   		OWF_Add_c.10:=OWF_Result[10].31;
   		OWF_Result[10].31:=0;
   		OWF_Result[11]:=OWF_Result[11] + 742245961+OWF_Add_c;
   		OWF_Add_c.11:=OWF_Result[11].31;
   		OWF_Result[11].31:=0;
   		OWF_Result[12]:=OWF_Result[12] + 1527470677+OWF_Add_c;
   		OWF_Add_c.12:=OWF_Result[12].31;
   		OWF_Result[12].31:=0;
   		OWF_Result[13]:=OWF_Result[13] + 104891933+OWF_Add_c;
   		OWF_Add_c.13:=OWF_Result[13].31;
   		OWF_Result[13].31:=0;
   		OWF_Result[14]:=OWF_Result[14] + 1414596320+OWF_Add_c;
   		OWF_Add_c.14:=OWF_Result[14].31;
   		OWF_Result[14].31:=0;
   		OWF_Result[15]:=OWF_Result[15] + 848151661+OWF_Add_c;
   		OWF_Add_c.15:=OWF_Result[15].31;
   		OWF_Result[15].31:=0;
   		OWF_Result[16]:=OWF_Result[16] + 1988122072+OWF_Add_c;
   		OWF_Add_c.16:=OWF_Result[16].31;
   		OWF_Result[16].31:=0;
   	End_If;
   	If OWF_Input[10].[29] Then
   		OWF_Result[0]:=OWF_Result[0] + 197995467+OWF_Add_c;
   		OWF_Add_c.0:=OWF_Result[0].31;
   		OWF_Result[0].31:=0;
   		OWF_Result[1]:=OWF_Result[1] + 1401962007+OWF_Add_c;
   		OWF_Add_c.1:=OWF_Result[1].31;
   		OWF_Result[1].31:=0;
   		OWF_Result[2]:=OWF_Result[2] + 1030218683+OWF_Add_c;
   		OWF_Add_c.2:=OWF_Result[2].31;
   		OWF_Result[2].31:=0;
   		OWF_Result[3]:=OWF_Result[3] + 1917186559+OWF_Add_c;
   		OWF_Add_c.3:=OWF_Result[3].31;
   		OWF_Result[3].31:=0;
   		OWF_Result[4]:=OWF_Result[4] + 1642815876+OWF_Add_c;
   		OWF_Add_c.4:=OWF_Result[4].31;
   		OWF_Result[4].31:=0;
   		OWF_Result[5]:=OWF_Result[5] + 126047613+OWF_Add_c;
   		OWF_Add_c.5:=OWF_Result[5].31;
   		OWF_Result[5].31:=0;
   		OWF_Result[6]:=OWF_Result[6] + 559790140+OWF_Add_c;
   		OWF_Add_c.6:=OWF_Result[6].31;
   		OWF_Result[6].31:=0;
   		OWF_Result[7]:=OWF_Result[7] + 2038093848+OWF_Add_c;
   		OWF_Add_c.7:=OWF_Result[7].31;
   		OWF_Result[7].31:=0;
   		OWF_Result[8]:=OWF_Result[8] + 221043685+OWF_Add_c;
   		OWF_Add_c.8:=OWF_Result[8].31;
   		OWF_Result[8].31:=0;
   		OWF_Result[9]:=OWF_Result[9] + 1671325631+OWF_Add_c;
   		OWF_Add_c.9:=OWF_Result[9].31;
   		OWF_Result[9].31:=0;
   		OWF_Result[10]:=OWF_Result[10] + 466139389+OWF_Add_c;
   		OWF_Add_c.10:=OWF_Result[10].31;
   		OWF_Result[10].31:=0;
   		OWF_Result[11]:=OWF_Result[11] + 25622731+OWF_Add_c;
   		OWF_Add_c.11:=OWF_Result[11].31;
   		OWF_Result[11].31:=0;
   		OWF_Result[12]:=OWF_Result[12] + 345868662+OWF_Add_c;
   		OWF_Add_c.12:=OWF_Result[12].31;
   		OWF_Result[12].31:=0;
   		OWF_Result[13]:=OWF_Result[13] + 822832112+OWF_Add_c;
   		OWF_Add_c.13:=OWF_Result[13].31;
   		OWF_Result[13].31:=0;
   		OWF_Result[14]:=OWF_Result[14] + 89551706+OWF_Add_c;
   		OWF_Add_c.14:=OWF_Result[14].31;
   		OWF_Result[14].31:=0;
   		OWF_Result[15]:=OWF_Result[15] + 1391211352+OWF_Add_c;
   		OWF_Add_c.15:=OWF_Result[15].31;
   		OWF_Result[15].31:=0;
   		OWF_Result[16]:=OWF_Result[16] + 1248625291+OWF_Add_c;
   		OWF_Add_c.16:=OWF_Result[16].31;
   		OWF_Result[16].31:=0;
   	End_If;
   	If OWF_Input[10].[30] Then
   		OWF_Result[0]:=OWF_Result[0] + 966732317+OWF_Add_c;
   		OWF_Add_c.0:=OWF_Result[0].31;
   		OWF_Result[0].31:=0;
   		OWF_Result[1]:=OWF_Result[1] + 1141530875+OWF_Add_c;
   		OWF_Add_c.1:=OWF_Result[1].31;
   		OWF_Result[1].31:=0;
   		OWF_Result[2]:=OWF_Result[2] + 1774163109+OWF_Add_c;
   		OWF_Add_c.2:=OWF_Result[2].31;
   		OWF_Result[2].31:=0;
   		OWF_Result[3]:=OWF_Result[3] + 1631047695+OWF_Add_c;
   		OWF_Add_c.3:=OWF_Result[3].31;
   		OWF_Result[3].31:=0;
   		OWF_Result[4]:=OWF_Result[4] + 1603525390+OWF_Add_c;
   		OWF_Add_c.4:=OWF_Result[4].31;
   		OWF_Result[4].31:=0;
   		OWF_Result[5]:=OWF_Result[5] + 626554573+OWF_Add_c;
   		OWF_Add_c.5:=OWF_Result[5].31;
   		OWF_Result[5].31:=0;
   		OWF_Result[6]:=OWF_Result[6] + 1641587637+OWF_Add_c;
   		OWF_Add_c.6:=OWF_Result[6].31;
   		OWF_Result[6].31:=0;
   		OWF_Result[7]:=OWF_Result[7] + 1028670148+OWF_Add_c;
   		OWF_Add_c.7:=OWF_Result[7].31;
   		OWF_Result[7].31:=0;
   		OWF_Result[8]:=OWF_Result[8] + 988622985+OWF_Add_c;
   		OWF_Add_c.8:=OWF_Result[8].31;
   		OWF_Result[8].31:=0;
   		OWF_Result[9]:=OWF_Result[9] + 1448454091+OWF_Add_c;
   		OWF_Add_c.9:=OWF_Result[9].31;
   		OWF_Result[9].31:=0;
   		OWF_Result[10]:=OWF_Result[10] + 532649595+OWF_Add_c;
   		OWF_Add_c.10:=OWF_Result[10].31;
   		OWF_Result[10].31:=0;
   		OWF_Result[11]:=OWF_Result[11] + 1443217515+OWF_Add_c;
   		OWF_Add_c.11:=OWF_Result[11].31;
   		OWF_Result[11].31:=0;
   		OWF_Result[12]:=OWF_Result[12] + 1792073364+OWF_Add_c;
   		OWF_Add_c.12:=OWF_Result[12].31;
   		OWF_Result[12].31:=0;
   		OWF_Result[13]:=OWF_Result[13] + 152898809+OWF_Add_c;
   		OWF_Add_c.13:=OWF_Result[13].31;
   		OWF_Result[13].31:=0;
   		OWF_Result[14]:=OWF_Result[14] + 354089137+OWF_Add_c;
   		OWF_Add_c.14:=OWF_Result[14].31;
   		OWF_Result[14].31:=0;
   		OWF_Result[15]:=OWF_Result[15] + 1049194702+OWF_Add_c;
   		OWF_Add_c.15:=OWF_Result[15].31;
   		OWF_Result[15].31:=0;
   		OWF_Result[16]:=OWF_Result[16] + 1707645884+OWF_Add_c;
   		OWF_Add_c.16:=OWF_Result[16].31;
   		OWF_Result[16].31:=0;
   	End_If;
   	If OWF_Input[10].[31] Then
   		OWF_Result[0]:=OWF_Result[0] + 1357392085+OWF_Add_c;
   		OWF_Add_c.0:=OWF_Result[0].31;
   		OWF_Result[0].31:=0;
   		OWF_Result[1]:=OWF_Result[1] + 130623031+OWF_Add_c;
   		OWF_Add_c.1:=OWF_Result[1].31;
   		OWF_Result[1].31:=0;
   		OWF_Result[2]:=OWF_Result[2] + 1002109794+OWF_Add_c;
   		OWF_Add_c.2:=OWF_Result[2].31;
   		OWF_Result[2].31:=0;
   		OWF_Result[3]:=OWF_Result[3] + 1001092841+OWF_Add_c;
   		OWF_Add_c.3:=OWF_Result[3].31;
   		OWF_Result[3].31:=0;
   		OWF_Result[4]:=OWF_Result[4] + 2057734046+OWF_Add_c;
   		OWF_Add_c.4:=OWF_Result[4].31;
   		OWF_Result[4].31:=0;
   		OWF_Result[5]:=OWF_Result[5] + 1800445178+OWF_Add_c;
   		OWF_Add_c.5:=OWF_Result[5].31;
   		OWF_Result[5].31:=0;
   		OWF_Result[6]:=OWF_Result[6] + 612634695+OWF_Add_c;
   		OWF_Add_c.6:=OWF_Result[6].31;
   		OWF_Result[6].31:=0;
   		OWF_Result[7]:=OWF_Result[7] + 25224326+OWF_Add_c;
   		OWF_Add_c.7:=OWF_Result[7].31;
   		OWF_Result[7].31:=0;
   		OWF_Result[8]:=OWF_Result[8] + 2106223567+OWF_Add_c;
   		OWF_Add_c.8:=OWF_Result[8].31;
   		OWF_Result[8].31:=0;
   		OWF_Result[9]:=OWF_Result[9] + 506405369+OWF_Add_c;
   		OWF_Add_c.9:=OWF_Result[9].31;
   		OWF_Result[9].31:=0;
   		OWF_Result[10]:=OWF_Result[10] + 1383246610+OWF_Add_c;
   		OWF_Add_c.10:=OWF_Result[10].31;
   		OWF_Result[10].31:=0;
   		OWF_Result[11]:=OWF_Result[11] + 2093993487+OWF_Add_c;
   		OWF_Add_c.11:=OWF_Result[11].31;
   		OWF_Result[11].31:=0;
   		OWF_Result[12]:=OWF_Result[12] + 338832249+OWF_Add_c;
   		OWF_Add_c.12:=OWF_Result[12].31;
   		OWF_Result[12].31:=0;
   		OWF_Result[13]:=OWF_Result[13] + 16899160+OWF_Add_c;
   		OWF_Add_c.13:=OWF_Result[13].31;
   		OWF_Result[13].31:=0;
   		OWF_Result[14]:=OWF_Result[14] + 1183329150+OWF_Add_c;
   		OWF_Add_c.14:=OWF_Result[14].31;
   		OWF_Result[14].31:=0;
   		OWF_Result[15]:=OWF_Result[15] + 505827814+OWF_Add_c;
   		OWF_Add_c.15:=OWF_Result[15].31;
   		OWF_Result[15].31:=0;
   		OWF_Result[16]:=OWF_Result[16] + 510585634+OWF_Add_c;
   		OWF_Add_c.16:=OWF_Result[16].31;
   		OWF_Result[16].31:=0;
   	End_If;
   	If OWF_Input[11].[0] Then
   		OWF_Result[0]:=OWF_Result[0] + 1007476166+OWF_Add_c;
   		OWF_Add_c.0:=OWF_Result[0].31;
   		OWF_Result[0].31:=0;
   		OWF_Result[1]:=OWF_Result[1] + 1504709985+OWF_Add_c;
   		OWF_Add_c.1:=OWF_Result[1].31;
   		OWF_Result[1].31:=0;
   		OWF_Result[2]:=OWF_Result[2] + 588918474+OWF_Add_c;
   		OWF_Add_c.2:=OWF_Result[2].31;
   		OWF_Result[2].31:=0;
   		OWF_Result[3]:=OWF_Result[3] + 1647627792+OWF_Add_c;
   		OWF_Add_c.3:=OWF_Result[3].31;
   		OWF_Result[3].31:=0;
   		OWF_Result[4]:=OWF_Result[4] + 1686612823+OWF_Add_c;
   		OWF_Add_c.4:=OWF_Result[4].31;
   		OWF_Result[4].31:=0;
   		OWF_Result[5]:=OWF_Result[5] + 1163719104+OWF_Add_c;
   		OWF_Add_c.5:=OWF_Result[5].31;
   		OWF_Result[5].31:=0;
   		OWF_Result[6]:=OWF_Result[6] + 127290704+OWF_Add_c;
   		OWF_Add_c.6:=OWF_Result[6].31;
   		OWF_Result[6].31:=0;
   		OWF_Result[7]:=OWF_Result[7] + 119227323+OWF_Add_c;
   		OWF_Add_c.7:=OWF_Result[7].31;
   		OWF_Result[7].31:=0;
   		OWF_Result[8]:=OWF_Result[8] + 2093562458+OWF_Add_c;
   		OWF_Add_c.8:=OWF_Result[8].31;
   		OWF_Result[8].31:=0;
   		OWF_Result[9]:=OWF_Result[9] + 1843045342+OWF_Add_c;
   		OWF_Add_c.9:=OWF_Result[9].31;
   		OWF_Result[9].31:=0;
   		OWF_Result[10]:=OWF_Result[10] + 2058220246+OWF_Add_c;
   		OWF_Add_c.10:=OWF_Result[10].31;
   		OWF_Result[10].31:=0;
   		OWF_Result[11]:=OWF_Result[11] + 1356791164+OWF_Add_c;
   		OWF_Add_c.11:=OWF_Result[11].31;
   		OWF_Result[11].31:=0;
   		OWF_Result[12]:=OWF_Result[12] + 853940386+OWF_Add_c;
   		OWF_Add_c.12:=OWF_Result[12].31;
   		OWF_Result[12].31:=0;
   		OWF_Result[13]:=OWF_Result[13] + 974030360+OWF_Add_c;
   		OWF_Add_c.13:=OWF_Result[13].31;
   		OWF_Result[13].31:=0;
   		OWF_Result[14]:=OWF_Result[14] + 1658027450+OWF_Add_c;
   		OWF_Add_c.14:=OWF_Result[14].31;
   		OWF_Result[14].31:=0;
   		OWF_Result[15]:=OWF_Result[15] + 1353014177+OWF_Add_c;
   		OWF_Add_c.15:=OWF_Result[15].31;
   		OWF_Result[15].31:=0;
   		OWF_Result[16]:=OWF_Result[16] + 149330334+OWF_Add_c;
   		OWF_Add_c.16:=OWF_Result[16].31;
   		OWF_Result[16].31:=0;
   	End_If;
   	If OWF_Input[11].[1] Then
   		OWF_Result[0]:=OWF_Result[0] + 1568466532+OWF_Add_c;
   		OWF_Add_c.0:=OWF_Result[0].31;
   		OWF_Result[0].31:=0;
   		OWF_Result[1]:=OWF_Result[1] + 1460316104+OWF_Add_c;
   		OWF_Add_c.1:=OWF_Result[1].31;
   		OWF_Result[1].31:=0;
   		OWF_Result[2]:=OWF_Result[2] + 1740708870+OWF_Add_c;
   		OWF_Add_c.2:=OWF_Result[2].31;
   		OWF_Result[2].31:=0;
   		OWF_Result[3]:=OWF_Result[3] + 339208175+OWF_Add_c;
   		OWF_Add_c.3:=OWF_Result[3].31;
   		OWF_Result[3].31:=0;
   		OWF_Result[4]:=OWF_Result[4] + 517379511+OWF_Add_c;
   		OWF_Add_c.4:=OWF_Result[4].31;
   		OWF_Result[4].31:=0;
   		OWF_Result[5]:=OWF_Result[5] + 864019991+OWF_Add_c;
   		OWF_Add_c.5:=OWF_Result[5].31;
   		OWF_Result[5].31:=0;
   		OWF_Result[6]:=OWF_Result[6] + 1026194771+OWF_Add_c;
   		OWF_Add_c.6:=OWF_Result[6].31;
   		OWF_Result[6].31:=0;
   		OWF_Result[7]:=OWF_Result[7] + 763406664+OWF_Add_c;
   		OWF_Add_c.7:=OWF_Result[7].31;
   		OWF_Result[7].31:=0;
   		OWF_Result[8]:=OWF_Result[8] + 1209552225+OWF_Add_c;
   		OWF_Add_c.8:=OWF_Result[8].31;
   		OWF_Result[8].31:=0;
   		OWF_Result[9]:=OWF_Result[9] + 1953270342+OWF_Add_c;
   		OWF_Add_c.9:=OWF_Result[9].31;
   		OWF_Result[9].31:=0;
   		OWF_Result[10]:=OWF_Result[10] + 934093539+OWF_Add_c;
   		OWF_Add_c.10:=OWF_Result[10].31;
   		OWF_Result[10].31:=0;
   		OWF_Result[11]:=OWF_Result[11] + 1096714606+OWF_Add_c;
   		OWF_Add_c.11:=OWF_Result[11].31;
   		OWF_Result[11].31:=0;
   		OWF_Result[12]:=OWF_Result[12] + 1321951524+OWF_Add_c;
   		OWF_Add_c.12:=OWF_Result[12].31;
   		OWF_Result[12].31:=0;
   		OWF_Result[13]:=OWF_Result[13] + 348944155+OWF_Add_c;
   		OWF_Add_c.13:=OWF_Result[13].31;
   		OWF_Result[13].31:=0;
   		OWF_Result[14]:=OWF_Result[14] + 1438305201+OWF_Add_c;
   		OWF_Add_c.14:=OWF_Result[14].31;
   		OWF_Result[14].31:=0;
   		OWF_Result[15]:=OWF_Result[15] + 30074938+OWF_Add_c;
   		OWF_Add_c.15:=OWF_Result[15].31;
   		OWF_Result[15].31:=0;
   		OWF_Result[16]:=OWF_Result[16] + 988811+OWF_Add_c;
   		OWF_Add_c.16:=OWF_Result[16].31;
   		OWF_Result[16].31:=0;
   	End_If;
   	If OWF_Input[11].[2] Then
   		OWF_Result[0]:=OWF_Result[0] + 1700235214+OWF_Add_c;
   		OWF_Add_c.0:=OWF_Result[0].31;
   		OWF_Result[0].31:=0;
   		OWF_Result[1]:=OWF_Result[1] + 831265880+OWF_Add_c;
   		OWF_Add_c.1:=OWF_Result[1].31;
   		OWF_Result[1].31:=0;
   		OWF_Result[2]:=OWF_Result[2] + 273999769+OWF_Add_c;
   		OWF_Add_c.2:=OWF_Result[2].31;
   		OWF_Result[2].31:=0;
   		OWF_Result[3]:=OWF_Result[3] + 999268093+OWF_Add_c;
   		OWF_Add_c.3:=OWF_Result[3].31;
   		OWF_Result[3].31:=0;
   		OWF_Result[4]:=OWF_Result[4] + 1123354466+OWF_Add_c;
   		OWF_Add_c.4:=OWF_Result[4].31;
   		OWF_Result[4].31:=0;
   		OWF_Result[5]:=OWF_Result[5] + 1328106541+OWF_Add_c;
   		OWF_Add_c.5:=OWF_Result[5].31;
   		OWF_Result[5].31:=0;
   		OWF_Result[6]:=OWF_Result[6] + 1723068716+OWF_Add_c;
   		OWF_Add_c.6:=OWF_Result[6].31;
   		OWF_Result[6].31:=0;
   		OWF_Result[7]:=OWF_Result[7] + 827383180+OWF_Add_c;
   		OWF_Add_c.7:=OWF_Result[7].31;
   		OWF_Result[7].31:=0;
   		OWF_Result[8]:=OWF_Result[8] + 531720932+OWF_Add_c;
   		OWF_Add_c.8:=OWF_Result[8].31;
   		OWF_Result[8].31:=0;
   		OWF_Result[9]:=OWF_Result[9] + 669468909+OWF_Add_c;
   		OWF_Add_c.9:=OWF_Result[9].31;
   		OWF_Result[9].31:=0;
   		OWF_Result[10]:=OWF_Result[10] + 923319981+OWF_Add_c;
   		OWF_Add_c.10:=OWF_Result[10].31;
   		OWF_Result[10].31:=0;
   		OWF_Result[11]:=OWF_Result[11] + 1373816862+OWF_Add_c;
   		OWF_Add_c.11:=OWF_Result[11].31;
   		OWF_Result[11].31:=0;
   		OWF_Result[12]:=OWF_Result[12] + 769977154+OWF_Add_c;
   		OWF_Add_c.12:=OWF_Result[12].31;
   		OWF_Result[12].31:=0;
   		OWF_Result[13]:=OWF_Result[13] + 812568572+OWF_Add_c;
   		OWF_Add_c.13:=OWF_Result[13].31;
   		OWF_Result[13].31:=0;
   		OWF_Result[14]:=OWF_Result[14] + 1928754765+OWF_Add_c;
   		OWF_Add_c.14:=OWF_Result[14].31;
   		OWF_Result[14].31:=0;
   		OWF_Result[15]:=OWF_Result[15] + 69475132+OWF_Add_c;
   		OWF_Add_c.15:=OWF_Result[15].31;
   		OWF_Result[15].31:=0;
   		OWF_Result[16]:=OWF_Result[16] + 327757708+OWF_Add_c;
   		OWF_Add_c.16:=OWF_Result[16].31;
   		OWF_Result[16].31:=0;
   	End_If;
   	If OWF_Input[11].[3] Then
   		OWF_Result[0]:=OWF_Result[0] + 1043167862+OWF_Add_c;
   		OWF_Add_c.0:=OWF_Result[0].31;
   		OWF_Result[0].31:=0;
   		OWF_Result[1]:=OWF_Result[1] + 1848703415+OWF_Add_c;
   		OWF_Add_c.1:=OWF_Result[1].31;
   		OWF_Result[1].31:=0;
   		OWF_Result[2]:=OWF_Result[2] + 503845072+OWF_Add_c;
   		OWF_Add_c.2:=OWF_Result[2].31;
   		OWF_Result[2].31:=0;
   		OWF_Result[3]:=OWF_Result[3] + 204900357+OWF_Add_c;
   		OWF_Add_c.3:=OWF_Result[3].31;
   		OWF_Result[3].31:=0;
   		OWF_Result[4]:=OWF_Result[4] + 2029563097+OWF_Add_c;
   		OWF_Add_c.4:=OWF_Result[4].31;
   		OWF_Result[4].31:=0;
   		OWF_Result[5]:=OWF_Result[5] + 1775074343+OWF_Add_c;
   		OWF_Add_c.5:=OWF_Result[5].31;
   		OWF_Result[5].31:=0;
   		OWF_Result[6]:=OWF_Result[6] + 341185552+OWF_Add_c;
   		OWF_Add_c.6:=OWF_Result[6].31;
   		OWF_Result[6].31:=0;
   		OWF_Result[7]:=OWF_Result[7] + 2120881534+OWF_Add_c;
   		OWF_Add_c.7:=OWF_Result[7].31;
   		OWF_Result[7].31:=0;
   		OWF_Result[8]:=OWF_Result[8] + 1527751763+OWF_Add_c;
   		OWF_Add_c.8:=OWF_Result[8].31;
   		OWF_Result[8].31:=0;
   		OWF_Result[9]:=OWF_Result[9] + 188765164+OWF_Add_c;
   		OWF_Add_c.9:=OWF_Result[9].31;
   		OWF_Result[9].31:=0;
   		OWF_Result[10]:=OWF_Result[10] + 1160032641+OWF_Add_c;
   		OWF_Add_c.10:=OWF_Result[10].31;
   		OWF_Result[10].31:=0;
   		OWF_Result[11]:=OWF_Result[11] + 645016819+OWF_Add_c;
   		OWF_Add_c.11:=OWF_Result[11].31;
   		OWF_Result[11].31:=0;
   		OWF_Result[12]:=OWF_Result[12] + 998595526+OWF_Add_c;
   		OWF_Add_c.12:=OWF_Result[12].31;
   		OWF_Result[12].31:=0;
   		OWF_Result[13]:=OWF_Result[13] + 1178367833+OWF_Add_c;
   		OWF_Add_c.13:=OWF_Result[13].31;
   		OWF_Result[13].31:=0;
   		OWF_Result[14]:=OWF_Result[14] + 2078383129+OWF_Add_c;
   		OWF_Add_c.14:=OWF_Result[14].31;
   		OWF_Result[14].31:=0;
   		OWF_Result[15]:=OWF_Result[15] + 1810699343+OWF_Add_c;
   		OWF_Add_c.15:=OWF_Result[15].31;
   		OWF_Result[15].31:=0;
   		OWF_Result[16]:=OWF_Result[16] + 1603179349+OWF_Add_c;
   		OWF_Add_c.16:=OWF_Result[16].31;
   		OWF_Result[16].31:=0;
   	End_If;
   	If OWF_Input[11].[4] Then
   		OWF_Result[0]:=OWF_Result[0] + 16774562+OWF_Add_c;
   		OWF_Add_c.0:=OWF_Result[0].31;
   		OWF_Result[0].31:=0;
   		OWF_Result[1]:=OWF_Result[1] + 1937203582+OWF_Add_c;
   		OWF_Add_c.1:=OWF_Result[1].31;
   		OWF_Result[1].31:=0;
   		OWF_Result[2]:=OWF_Result[2] + 2141651730+OWF_Add_c;
   		OWF_Add_c.2:=OWF_Result[2].31;
   		OWF_Result[2].31:=0;
   		OWF_Result[3]:=OWF_Result[3] + 123641449+OWF_Add_c;
   		OWF_Add_c.3:=OWF_Result[3].31;
   		OWF_Result[3].31:=0;
   		OWF_Result[4]:=OWF_Result[4] + 1249486137+OWF_Add_c;
   		OWF_Add_c.4:=OWF_Result[4].31;
   		OWF_Result[4].31:=0;
   		OWF_Result[5]:=OWF_Result[5] + 1761614983+OWF_Add_c;
   		OWF_Add_c.5:=OWF_Result[5].31;
   		OWF_Result[5].31:=0;
   		OWF_Result[6]:=OWF_Result[6] + 1524506566+OWF_Add_c;
   		OWF_Add_c.6:=OWF_Result[6].31;
   		OWF_Result[6].31:=0;
   		OWF_Result[7]:=OWF_Result[7] + 1674479690+OWF_Add_c;
   		OWF_Add_c.7:=OWF_Result[7].31;
   		OWF_Result[7].31:=0;
   		OWF_Result[8]:=OWF_Result[8] + 1781150491+OWF_Add_c;
   		OWF_Add_c.8:=OWF_Result[8].31;
   		OWF_Result[8].31:=0;
   		OWF_Result[9]:=OWF_Result[9] + 1077235569+OWF_Add_c;
   		OWF_Add_c.9:=OWF_Result[9].31;
   		OWF_Result[9].31:=0;
   		OWF_Result[10]:=OWF_Result[10] + 906319697+OWF_Add_c;
   		OWF_Add_c.10:=OWF_Result[10].31;
   		OWF_Result[10].31:=0;
   		OWF_Result[11]:=OWF_Result[11] + 1482044083+OWF_Add_c;
   		OWF_Add_c.11:=OWF_Result[11].31;
   		OWF_Result[11].31:=0;
   		OWF_Result[12]:=OWF_Result[12] + 1323002605+OWF_Add_c;
   		OWF_Add_c.12:=OWF_Result[12].31;
   		OWF_Result[12].31:=0;
   		OWF_Result[13]:=OWF_Result[13] + 1102385938+OWF_Add_c;
   		OWF_Add_c.13:=OWF_Result[13].31;
   		OWF_Result[13].31:=0;
   		OWF_Result[14]:=OWF_Result[14] + 1043072459+OWF_Add_c;
   		OWF_Add_c.14:=OWF_Result[14].31;
   		OWF_Result[14].31:=0;
   		OWF_Result[15]:=OWF_Result[15] + 1279231835+OWF_Add_c;
   		OWF_Add_c.15:=OWF_Result[15].31;
   		OWF_Result[15].31:=0;
   		OWF_Result[16]:=OWF_Result[16] + 881943477+OWF_Add_c;
   		OWF_Add_c.16:=OWF_Result[16].31;
   		OWF_Result[16].31:=0;
   	End_If;
   	If OWF_Input[11].[5] Then
   		OWF_Result[0]:=OWF_Result[0] + 1185323519+OWF_Add_c;
   		OWF_Add_c.0:=OWF_Result[0].31;
   		OWF_Result[0].31:=0;
   		OWF_Result[1]:=OWF_Result[1] + 1959708271+OWF_Add_c;
   		OWF_Add_c.1:=OWF_Result[1].31;
   		OWF_Result[1].31:=0;
   		OWF_Result[2]:=OWF_Result[2] + 1001251338+OWF_Add_c;
   		OWF_Add_c.2:=OWF_Result[2].31;
   		OWF_Result[2].31:=0;
   		OWF_Result[3]:=OWF_Result[3] + 1077039075+OWF_Add_c;
   		OWF_Add_c.3:=OWF_Result[3].31;
   		OWF_Result[3].31:=0;
   		OWF_Result[4]:=OWF_Result[4] + 912657761+OWF_Add_c;
   		OWF_Add_c.4:=OWF_Result[4].31;
   		OWF_Result[4].31:=0;
   		OWF_Result[5]:=OWF_Result[5] + 1566133902+OWF_Add_c;
   		OWF_Add_c.5:=OWF_Result[5].31;
   		OWF_Result[5].31:=0;
   		OWF_Result[6]:=OWF_Result[6] + 2079545881+OWF_Add_c;
   		OWF_Add_c.6:=OWF_Result[6].31;
   		OWF_Result[6].31:=0;
   		OWF_Result[7]:=OWF_Result[7] + 1492050917+OWF_Add_c;
   		OWF_Add_c.7:=OWF_Result[7].31;
   		OWF_Result[7].31:=0;
   		OWF_Result[8]:=OWF_Result[8] + 1277398732+OWF_Add_c;
   		OWF_Add_c.8:=OWF_Result[8].31;
   		OWF_Result[8].31:=0;
   		OWF_Result[9]:=OWF_Result[9] + 438901726+OWF_Add_c;
   		OWF_Add_c.9:=OWF_Result[9].31;
   		OWF_Result[9].31:=0;
   		OWF_Result[10]:=OWF_Result[10] + 711557165+OWF_Add_c;
   		OWF_Add_c.10:=OWF_Result[10].31;
   		OWF_Result[10].31:=0;
   		OWF_Result[11]:=OWF_Result[11] + 1022238460+OWF_Add_c;
   		OWF_Add_c.11:=OWF_Result[11].31;
   		OWF_Result[11].31:=0;
   		OWF_Result[12]:=OWF_Result[12] + 370384684+OWF_Add_c;
   		OWF_Add_c.12:=OWF_Result[12].31;
   		OWF_Result[12].31:=0;
   		OWF_Result[13]:=OWF_Result[13] + 984834140+OWF_Add_c;
   		OWF_Add_c.13:=OWF_Result[13].31;
   		OWF_Result[13].31:=0;
   		OWF_Result[14]:=OWF_Result[14] + 1324280833+OWF_Add_c;
   		OWF_Add_c.14:=OWF_Result[14].31;
   		OWF_Result[14].31:=0;
   		OWF_Result[15]:=OWF_Result[15] + 1223498052+OWF_Add_c;
   		OWF_Add_c.15:=OWF_Result[15].31;
   		OWF_Result[15].31:=0;
   		OWF_Result[16]:=OWF_Result[16] + 541972467+OWF_Add_c;
   		OWF_Add_c.16:=OWF_Result[16].31;
   		OWF_Result[16].31:=0;
   	End_If;
   	If OWF_Input[11].[6] Then
   		OWF_Result[0]:=OWF_Result[0] + 1162786490+OWF_Add_c;
   		OWF_Add_c.0:=OWF_Result[0].31;
   		OWF_Result[0].31:=0;
   		OWF_Result[1]:=OWF_Result[1] + 126987719+OWF_Add_c;
   		OWF_Add_c.1:=OWF_Result[1].31;
   		OWF_Result[1].31:=0;
   		OWF_Result[2]:=OWF_Result[2] + 171798537+OWF_Add_c;
   		OWF_Add_c.2:=OWF_Result[2].31;
   		OWF_Result[2].31:=0;
   		OWF_Result[3]:=OWF_Result[3] + 1671423715+OWF_Add_c;
   		OWF_Add_c.3:=OWF_Result[3].31;
   		OWF_Result[3].31:=0;
   		OWF_Result[4]:=OWF_Result[4] + 126324653+OWF_Add_c;
   		OWF_Add_c.4:=OWF_Result[4].31;
   		OWF_Result[4].31:=0;
   		OWF_Result[5]:=OWF_Result[5] + 1359613574+OWF_Add_c;
   		OWF_Add_c.5:=OWF_Result[5].31;
   		OWF_Result[5].31:=0;
   		OWF_Result[6]:=OWF_Result[6] + 1153736861+OWF_Add_c;
   		OWF_Add_c.6:=OWF_Result[6].31;
   		OWF_Result[6].31:=0;
   		OWF_Result[7]:=OWF_Result[7] + 1791938875+OWF_Add_c;
   		OWF_Add_c.7:=OWF_Result[7].31;
   		OWF_Result[7].31:=0;
   		OWF_Result[8]:=OWF_Result[8] + 917211193+OWF_Add_c;
   		OWF_Add_c.8:=OWF_Result[8].31;
   		OWF_Result[8].31:=0;
   		OWF_Result[9]:=OWF_Result[9] + 1408684390+OWF_Add_c;
   		OWF_Add_c.9:=OWF_Result[9].31;
   		OWF_Result[9].31:=0;
   		OWF_Result[10]:=OWF_Result[10] + 844894848+OWF_Add_c;
   		OWF_Add_c.10:=OWF_Result[10].31;
   		OWF_Result[10].31:=0;
   		OWF_Result[11]:=OWF_Result[11] + 1669965479+OWF_Add_c;
   		OWF_Add_c.11:=OWF_Result[11].31;
   		OWF_Result[11].31:=0;
   		OWF_Result[12]:=OWF_Result[12] + 163113283+OWF_Add_c;
   		OWF_Add_c.12:=OWF_Result[12].31;
   		OWF_Result[12].31:=0;
   		OWF_Result[13]:=OWF_Result[13] + 626528550+OWF_Add_c;
   		OWF_Add_c.13:=OWF_Result[13].31;
   		OWF_Result[13].31:=0;
   		OWF_Result[14]:=OWF_Result[14] + 589313573+OWF_Add_c;
   		OWF_Add_c.14:=OWF_Result[14].31;
   		OWF_Result[14].31:=0;
   		OWF_Result[15]:=OWF_Result[15] + 1610018817+OWF_Add_c;
   		OWF_Add_c.15:=OWF_Result[15].31;
   		OWF_Result[15].31:=0;
   		OWF_Result[16]:=OWF_Result[16] + 444635992+OWF_Add_c;
   		OWF_Add_c.16:=OWF_Result[16].31;
   		OWF_Result[16].31:=0;
   	End_If;
   	If OWF_Input[11].[7] Then
   		OWF_Result[0]:=OWF_Result[0] + 238660872+OWF_Add_c;
   		OWF_Add_c.0:=OWF_Result[0].31;
   		OWF_Result[0].31:=0;
   		OWF_Result[1]:=OWF_Result[1] + 1205386123+OWF_Add_c;
   		OWF_Add_c.1:=OWF_Result[1].31;
   		OWF_Result[1].31:=0;
   		OWF_Result[2]:=OWF_Result[2] + 745841071+OWF_Add_c;
   		OWF_Add_c.2:=OWF_Result[2].31;
   		OWF_Result[2].31:=0;
   		OWF_Result[3]:=OWF_Result[3] + 687757852+OWF_Add_c;
   		OWF_Add_c.3:=OWF_Result[3].31;
   		OWF_Result[3].31:=0;
   		OWF_Result[4]:=OWF_Result[4] + 2009189753+OWF_Add_c;
   		OWF_Add_c.4:=OWF_Result[4].31;
   		OWF_Result[4].31:=0;
   		OWF_Result[5]:=OWF_Result[5] + 1740287639+OWF_Add_c;
   		OWF_Add_c.5:=OWF_Result[5].31;
   		OWF_Result[5].31:=0;
   		OWF_Result[6]:=OWF_Result[6] + 249867650+OWF_Add_c;
   		OWF_Add_c.6:=OWF_Result[6].31;
   		OWF_Result[6].31:=0;
   		OWF_Result[7]:=OWF_Result[7] + 691165392+OWF_Add_c;
   		OWF_Add_c.7:=OWF_Result[7].31;
   		OWF_Result[7].31:=0;
   		OWF_Result[8]:=OWF_Result[8] + 415030103+OWF_Add_c;
   		OWF_Add_c.8:=OWF_Result[8].31;
   		OWF_Result[8].31:=0;
   		OWF_Result[9]:=OWF_Result[9] + 1869752015+OWF_Add_c;
   		OWF_Add_c.9:=OWF_Result[9].31;
   		OWF_Result[9].31:=0;
   		OWF_Result[10]:=OWF_Result[10] + 422860613+OWF_Add_c;
   		OWF_Add_c.10:=OWF_Result[10].31;
   		OWF_Result[10].31:=0;
   		OWF_Result[11]:=OWF_Result[11] + 2089779412+OWF_Add_c;
   		OWF_Add_c.11:=OWF_Result[11].31;
   		OWF_Result[11].31:=0;
   		OWF_Result[12]:=OWF_Result[12] + 626521711+OWF_Add_c;
   		OWF_Add_c.12:=OWF_Result[12].31;
   		OWF_Result[12].31:=0;
   		OWF_Result[13]:=OWF_Result[13] + 523975610+OWF_Add_c;
   		OWF_Add_c.13:=OWF_Result[13].31;
   		OWF_Result[13].31:=0;
   		OWF_Result[14]:=OWF_Result[14] + 1085416245+OWF_Add_c;
   		OWF_Add_c.14:=OWF_Result[14].31;
   		OWF_Result[14].31:=0;
   		OWF_Result[15]:=OWF_Result[15] + 662822616+OWF_Add_c;
   		OWF_Add_c.15:=OWF_Result[15].31;
   		OWF_Result[15].31:=0;
   		OWF_Result[16]:=OWF_Result[16] + 1982964767+OWF_Add_c;
   		OWF_Add_c.16:=OWF_Result[16].31;
   		OWF_Result[16].31:=0;
   	End_If;
   	If OWF_Input[11].[8] Then
   		OWF_Result[0]:=OWF_Result[0] + 1147887739+OWF_Add_c;
   		OWF_Add_c.0:=OWF_Result[0].31;
   		OWF_Result[0].31:=0;
   		OWF_Result[1]:=OWF_Result[1] + 670270591+OWF_Add_c;
   		OWF_Add_c.1:=OWF_Result[1].31;
   		OWF_Result[1].31:=0;
   		OWF_Result[2]:=OWF_Result[2] + 1918427275+OWF_Add_c;
   		OWF_Add_c.2:=OWF_Result[2].31;
   		OWF_Result[2].31:=0;
   		OWF_Result[3]:=OWF_Result[3] + 1192408481+OWF_Add_c;
   		OWF_Add_c.3:=OWF_Result[3].31;
   		OWF_Result[3].31:=0;
   		OWF_Result[4]:=OWF_Result[4] + 138457706+OWF_Add_c;
   		OWF_Add_c.4:=OWF_Result[4].31;
   		OWF_Result[4].31:=0;
   		OWF_Result[5]:=OWF_Result[5] + 347687872+OWF_Add_c;
   		OWF_Add_c.5:=OWF_Result[5].31;
   		OWF_Result[5].31:=0;
   		OWF_Result[6]:=OWF_Result[6] + 231537152+OWF_Add_c;
   		OWF_Add_c.6:=OWF_Result[6].31;
   		OWF_Result[6].31:=0;
   		OWF_Result[7]:=OWF_Result[7] + 603699292+OWF_Add_c;
   		OWF_Add_c.7:=OWF_Result[7].31;
   		OWF_Result[7].31:=0;
   		OWF_Result[8]:=OWF_Result[8] + 672706039+OWF_Add_c;
   		OWF_Add_c.8:=OWF_Result[8].31;
   		OWF_Result[8].31:=0;
   		OWF_Result[9]:=OWF_Result[9] + 213476514+OWF_Add_c;
   		OWF_Add_c.9:=OWF_Result[9].31;
   		OWF_Result[9].31:=0;
   		OWF_Result[10]:=OWF_Result[10] + 1301300293+OWF_Add_c;
   		OWF_Add_c.10:=OWF_Result[10].31;
   		OWF_Result[10].31:=0;
   		OWF_Result[11]:=OWF_Result[11] + 1650338655+OWF_Add_c;
   		OWF_Add_c.11:=OWF_Result[11].31;
   		OWF_Result[11].31:=0;
   		OWF_Result[12]:=OWF_Result[12] + 800302141+OWF_Add_c;
   		OWF_Add_c.12:=OWF_Result[12].31;
   		OWF_Result[12].31:=0;
   		OWF_Result[13]:=OWF_Result[13] + 255254240+OWF_Add_c;
   		OWF_Add_c.13:=OWF_Result[13].31;
   		OWF_Result[13].31:=0;
   		OWF_Result[14]:=OWF_Result[14] + 1933455758+OWF_Add_c;
   		OWF_Add_c.14:=OWF_Result[14].31;
   		OWF_Result[14].31:=0;
   		OWF_Result[15]:=OWF_Result[15] + 736844305+OWF_Add_c;
   		OWF_Add_c.15:=OWF_Result[15].31;
   		OWF_Result[15].31:=0;
   		OWF_Result[16]:=OWF_Result[16] + 1841703559+OWF_Add_c;
   		OWF_Add_c.16:=OWF_Result[16].31;
   		OWF_Result[16].31:=0;
   	End_If;
   	If OWF_Input[11].[9] Then
   		OWF_Result[0]:=OWF_Result[0] + 653311066+OWF_Add_c;
   		OWF_Add_c.0:=OWF_Result[0].31;
   		OWF_Result[0].31:=0;
   		OWF_Result[1]:=OWF_Result[1] + 13547699+OWF_Add_c;
   		OWF_Add_c.1:=OWF_Result[1].31;
   		OWF_Result[1].31:=0;
   		OWF_Result[2]:=OWF_Result[2] + 838482689+OWF_Add_c;
   		OWF_Add_c.2:=OWF_Result[2].31;
   		OWF_Result[2].31:=0;
   		OWF_Result[3]:=OWF_Result[3] + 1006972684+OWF_Add_c;
   		OWF_Add_c.3:=OWF_Result[3].31;
   		OWF_Result[3].31:=0;
   		OWF_Result[4]:=OWF_Result[4] + 328883471+OWF_Add_c;
   		OWF_Add_c.4:=OWF_Result[4].31;
   		OWF_Result[4].31:=0;
   		OWF_Result[5]:=OWF_Result[5] + 1080319626+OWF_Add_c;
   		OWF_Add_c.5:=OWF_Result[5].31;
   		OWF_Result[5].31:=0;
   		OWF_Result[6]:=OWF_Result[6] + 731358565+OWF_Add_c;
   		OWF_Add_c.6:=OWF_Result[6].31;
   		OWF_Result[6].31:=0;
   		OWF_Result[7]:=OWF_Result[7] + 945543794+OWF_Add_c;
   		OWF_Add_c.7:=OWF_Result[7].31;
   		OWF_Result[7].31:=0;
   		OWF_Result[8]:=OWF_Result[8] + 1295547745+OWF_Add_c;
   		OWF_Add_c.8:=OWF_Result[8].31;
   		OWF_Result[8].31:=0;
   		OWF_Result[9]:=OWF_Result[9] + 31813743+OWF_Add_c;
   		OWF_Add_c.9:=OWF_Result[9].31;
   		OWF_Result[9].31:=0;
   		OWF_Result[10]:=OWF_Result[10] + 1261015854+OWF_Add_c;
   		OWF_Add_c.10:=OWF_Result[10].31;
   		OWF_Result[10].31:=0;
   		OWF_Result[11]:=OWF_Result[11] + 1410311323+OWF_Add_c;
   		OWF_Add_c.11:=OWF_Result[11].31;
   		OWF_Result[11].31:=0;
   		OWF_Result[12]:=OWF_Result[12] + 2128158986+OWF_Add_c;
   		OWF_Add_c.12:=OWF_Result[12].31;
   		OWF_Result[12].31:=0;
   		OWF_Result[13]:=OWF_Result[13] + 1912178265+OWF_Add_c;
   		OWF_Add_c.13:=OWF_Result[13].31;
   		OWF_Result[13].31:=0;
   		OWF_Result[14]:=OWF_Result[14] + 2077338334+OWF_Add_c;
   		OWF_Add_c.14:=OWF_Result[14].31;
   		OWF_Result[14].31:=0;
   		OWF_Result[15]:=OWF_Result[15] + 1398427904+OWF_Add_c;
   		OWF_Add_c.15:=OWF_Result[15].31;
   		OWF_Result[15].31:=0;
   		OWF_Result[16]:=OWF_Result[16] + 918416271+OWF_Add_c;
   		OWF_Add_c.16:=OWF_Result[16].31;
   		OWF_Result[16].31:=0;
   	End_If;
   	If OWF_Input[11].[10] Then
   		OWF_Result[0]:=OWF_Result[0] + 1667652198+OWF_Add_c;
   		OWF_Add_c.0:=OWF_Result[0].31;
   		OWF_Result[0].31:=0;
   		OWF_Result[1]:=OWF_Result[1] + 1571001387+OWF_Add_c;
   		OWF_Add_c.1:=OWF_Result[1].31;
   		OWF_Result[1].31:=0;
   		OWF_Result[2]:=OWF_Result[2] + 535742622+OWF_Add_c;
   		OWF_Add_c.2:=OWF_Result[2].31;
   		OWF_Result[2].31:=0;
   		OWF_Result[3]:=OWF_Result[3] + 1270090821+OWF_Add_c;
   		OWF_Add_c.3:=OWF_Result[3].31;
   		OWF_Result[3].31:=0;
   		OWF_Result[4]:=OWF_Result[4] + 1553530389+OWF_Add_c;
   		OWF_Add_c.4:=OWF_Result[4].31;
   		OWF_Result[4].31:=0;
   		OWF_Result[5]:=OWF_Result[5] + 2042097332+OWF_Add_c;
   		OWF_Add_c.5:=OWF_Result[5].31;
   		OWF_Result[5].31:=0;
   		OWF_Result[6]:=OWF_Result[6] + 2017684049+OWF_Add_c;
   		OWF_Add_c.6:=OWF_Result[6].31;
   		OWF_Result[6].31:=0;
   		OWF_Result[7]:=OWF_Result[7] + 2128486148+OWF_Add_c;
   		OWF_Add_c.7:=OWF_Result[7].31;
   		OWF_Result[7].31:=0;
   		OWF_Result[8]:=OWF_Result[8] + 1132700769+OWF_Add_c;
   		OWF_Add_c.8:=OWF_Result[8].31;
   		OWF_Result[8].31:=0;
   		OWF_Result[9]:=OWF_Result[9] + 1333860019+OWF_Add_c;
   		OWF_Add_c.9:=OWF_Result[9].31;
   		OWF_Result[9].31:=0;
   		OWF_Result[10]:=OWF_Result[10] + 1111911107+OWF_Add_c;
   		OWF_Add_c.10:=OWF_Result[10].31;
   		OWF_Result[10].31:=0;
   		OWF_Result[11]:=OWF_Result[11] + 1993892775+OWF_Add_c;
   		OWF_Add_c.11:=OWF_Result[11].31;
   		OWF_Result[11].31:=0;
   		OWF_Result[12]:=OWF_Result[12] + 540831246+OWF_Add_c;
   		OWF_Add_c.12:=OWF_Result[12].31;
   		OWF_Result[12].31:=0;
   		OWF_Result[13]:=OWF_Result[13] + 913455896+OWF_Add_c;
   		OWF_Add_c.13:=OWF_Result[13].31;
   		OWF_Result[13].31:=0;
   		OWF_Result[14]:=OWF_Result[14] + 796372115+OWF_Add_c;
   		OWF_Add_c.14:=OWF_Result[14].31;
   		OWF_Result[14].31:=0;
   		OWF_Result[15]:=OWF_Result[15] + 1207639928+OWF_Add_c;
   		OWF_Add_c.15:=OWF_Result[15].31;
   		OWF_Result[15].31:=0;
   		OWF_Result[16]:=OWF_Result[16] + 354716243+OWF_Add_c;
   		OWF_Add_c.16:=OWF_Result[16].31;
   		OWF_Result[16].31:=0;
   	End_If;
   	If OWF_Input[11].[11] Then
   		OWF_Result[0]:=OWF_Result[0] + 443861865+OWF_Add_c;
   		OWF_Add_c.0:=OWF_Result[0].31;
   		OWF_Result[0].31:=0;
   		OWF_Result[1]:=OWF_Result[1] + 1063977421+OWF_Add_c;
   		OWF_Add_c.1:=OWF_Result[1].31;
   		OWF_Result[1].31:=0;
   		OWF_Result[2]:=OWF_Result[2] + 1006340556+OWF_Add_c;
   		OWF_Add_c.2:=OWF_Result[2].31;
   		OWF_Result[2].31:=0;
   		OWF_Result[3]:=OWF_Result[3] + 1972055115+OWF_Add_c;
   		OWF_Add_c.3:=OWF_Result[3].31;
   		OWF_Result[3].31:=0;
   		OWF_Result[4]:=OWF_Result[4] + 615966915+OWF_Add_c;
   		OWF_Add_c.4:=OWF_Result[4].31;
   		OWF_Result[4].31:=0;
   		OWF_Result[5]:=OWF_Result[5] + 836753688+OWF_Add_c;
   		OWF_Add_c.5:=OWF_Result[5].31;
   		OWF_Result[5].31:=0;
   		OWF_Result[6]:=OWF_Result[6] + 1549512770+OWF_Add_c;
   		OWF_Add_c.6:=OWF_Result[6].31;
   		OWF_Result[6].31:=0;
   		OWF_Result[7]:=OWF_Result[7] + 1134835744+OWF_Add_c;
   		OWF_Add_c.7:=OWF_Result[7].31;
   		OWF_Result[7].31:=0;
   		OWF_Result[8]:=OWF_Result[8] + 639600176+OWF_Add_c;
   		OWF_Add_c.8:=OWF_Result[8].31;
   		OWF_Result[8].31:=0;
   		OWF_Result[9]:=OWF_Result[9] + 1887339535+OWF_Add_c;
   		OWF_Add_c.9:=OWF_Result[9].31;
   		OWF_Result[9].31:=0;
   		OWF_Result[10]:=OWF_Result[10] + 2104225157+OWF_Add_c;
   		OWF_Add_c.10:=OWF_Result[10].31;
   		OWF_Result[10].31:=0;
   		OWF_Result[11]:=OWF_Result[11] + 1224171535+OWF_Add_c;
   		OWF_Add_c.11:=OWF_Result[11].31;
   		OWF_Result[11].31:=0;
   		OWF_Result[12]:=OWF_Result[12] + 2025775365+OWF_Add_c;
   		OWF_Add_c.12:=OWF_Result[12].31;
   		OWF_Result[12].31:=0;
   		OWF_Result[13]:=OWF_Result[13] + 321398187+OWF_Add_c;
   		OWF_Add_c.13:=OWF_Result[13].31;
   		OWF_Result[13].31:=0;
   		OWF_Result[14]:=OWF_Result[14] + 477405553+OWF_Add_c;
   		OWF_Add_c.14:=OWF_Result[14].31;
   		OWF_Result[14].31:=0;
   		OWF_Result[15]:=OWF_Result[15] + 1083910466+OWF_Add_c;
   		OWF_Add_c.15:=OWF_Result[15].31;
   		OWF_Result[15].31:=0;
   		OWF_Result[16]:=OWF_Result[16] + 729656794+OWF_Add_c;
   		OWF_Add_c.16:=OWF_Result[16].31;
   		OWF_Result[16].31:=0;
   	End_If;
   	If OWF_Input[11].[12] Then
   		OWF_Result[0]:=OWF_Result[0] + 1612392199+OWF_Add_c;
   		OWF_Add_c.0:=OWF_Result[0].31;
   		OWF_Result[0].31:=0;
   		OWF_Result[1]:=OWF_Result[1] + 479243269+OWF_Add_c;
   		OWF_Add_c.1:=OWF_Result[1].31;
   		OWF_Result[1].31:=0;
   		OWF_Result[2]:=OWF_Result[2] + 867278740+OWF_Add_c;
   		OWF_Add_c.2:=OWF_Result[2].31;
   		OWF_Result[2].31:=0;
   		OWF_Result[3]:=OWF_Result[3] + 1518275338+OWF_Add_c;
   		OWF_Add_c.3:=OWF_Result[3].31;
   		OWF_Result[3].31:=0;
   		OWF_Result[4]:=OWF_Result[4] + 575766006+OWF_Add_c;
   		OWF_Add_c.4:=OWF_Result[4].31;
